   "ALARM_PT402" := ("PT402_VAL" > "PT402_HIGH") OR ("ALARM_PT402" AND NOT #CLEAR);
   "ALARM_PT501" := ("PT501_VAL" < "PT501_LOW_C") OR ("ALARM_PT501" AND NOT #CLEAR);
   "ALARM_PT502" := ("PT502_VAL" > "PT502_HIGH") OR ("ALARM_PT502" AND NOT #CLEAR);
   "ALARM_PT601" := ("PT601_VAL" >= "PT601_HIGH") OR ("ALARM_PT601" AND NOT #CLEAR);
   "ALARM_PT801" := ("PT801_VAL" < "PT801_LOW") OR ("ALARM_PT801" AND NOT #CLEAR);
   "ALARM_PT901" := ("PT901_VAL" > "PT901_HIGH") OR ("ALARM_PT901" AND NOT #CLEAR);
   "ALARM_DOORS_OPEN" := NOT "ABORT_ON" AND NOT "STEP_0_ON" AND NOT "DOORS_CLOSED" AND "AlwaysFALSE";
END_REGION

REGION Network 2
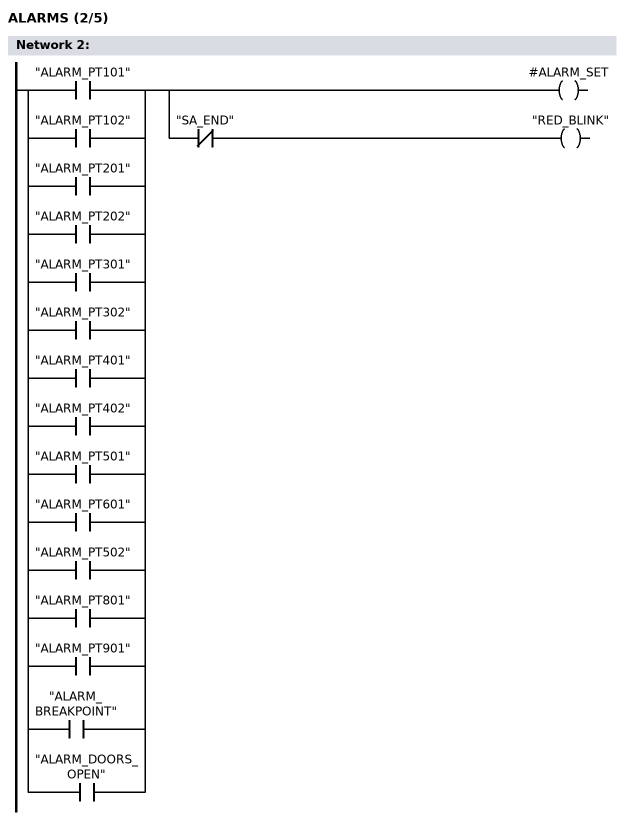
   RUNG wire#powerrail
      Contact( "ALARM_PT101" )
      wire#w1
      Coil( #ALARM_SET )
   END_RUNG
   RUNG wire#powerrail
      Contact( "ALARM_PT102" )
   END_RUNG wire#w1
   RUNG wire#powerrail
      Contact( "ALARM_PT201" )
   END_RUNG wire#w1
   RUNG wire#powerrail
      Contact( "ALARM_PT202" )
   END_RUNG wire#w1
   RUNG wire#powerrail
      Contact( "ALARM_PT301" )
   END_RUNG wire#w1
   RUNG wire#powerrail
      Contact( "ALARM_PT302" )
   END_RUNG wire#w1
   RUNG wire#powerrail
      Contact( "ALARM_PT401" )
   END_RUNG wire#w1
   RUNG wire#powerrail
      Contact( "ALARM_PT402" )
   END_RUNG wire#w1
   RUNG wire#powerrail
      Contact( "ALARM_PT501" )
   END_RUNG wire#w1
   RUNG wire#powerrail
      Contact( "ALARM_PT601" )
   END_RUNG wire#w1
   RUNG wire#powerrail
      Contact( "ALARM_PT502" )
   END_RUNG wire#w1
   RUNG wire#powerrail
      Contact( "ALARM_PT801" )
   END_RUNG wire#w1
   RUNG wire#powerrail
      Contact( "ALARM_PT901" )
   END_RUNG wire#w1
   RUNG wire#powerrail
      Contact( "ALARM_BREAKPOINT" )
   END_RUNG wire#w1
   RUNG wire#powerrail
      Contact( "ALARM_DOORS_OPEN" )
   END_RUNG wire#w1
   RUNG wire#w1
      I_Contact( "SA_END" )
      Coil( "RED_BLINK" )
   END_RUNG
   // the same network as SCL:
   #ALARM_SET := "ALARM_PT101" OR "ALARM_PT102" OR "ALARM_PT201" OR "ALARM_PT202" OR "ALARM_PT301" OR "ALARM_PT302" OR "ALARM_PT401" OR "ALARM_PT402" OR "ALARM_PT501" OR "ALARM_PT601" OR "ALARM_PT502" OR "ALARM_PT801" OR "ALARM_PT901" OR "ALARM_BREAKPOINT" OR "ALARM_DOORS_OPEN";
   "RED_BLINK" := #ALARM_SET AND NOT "SA_END";
END_REGION

REGION Network 3
   // PV701 Limit Switch Alarm
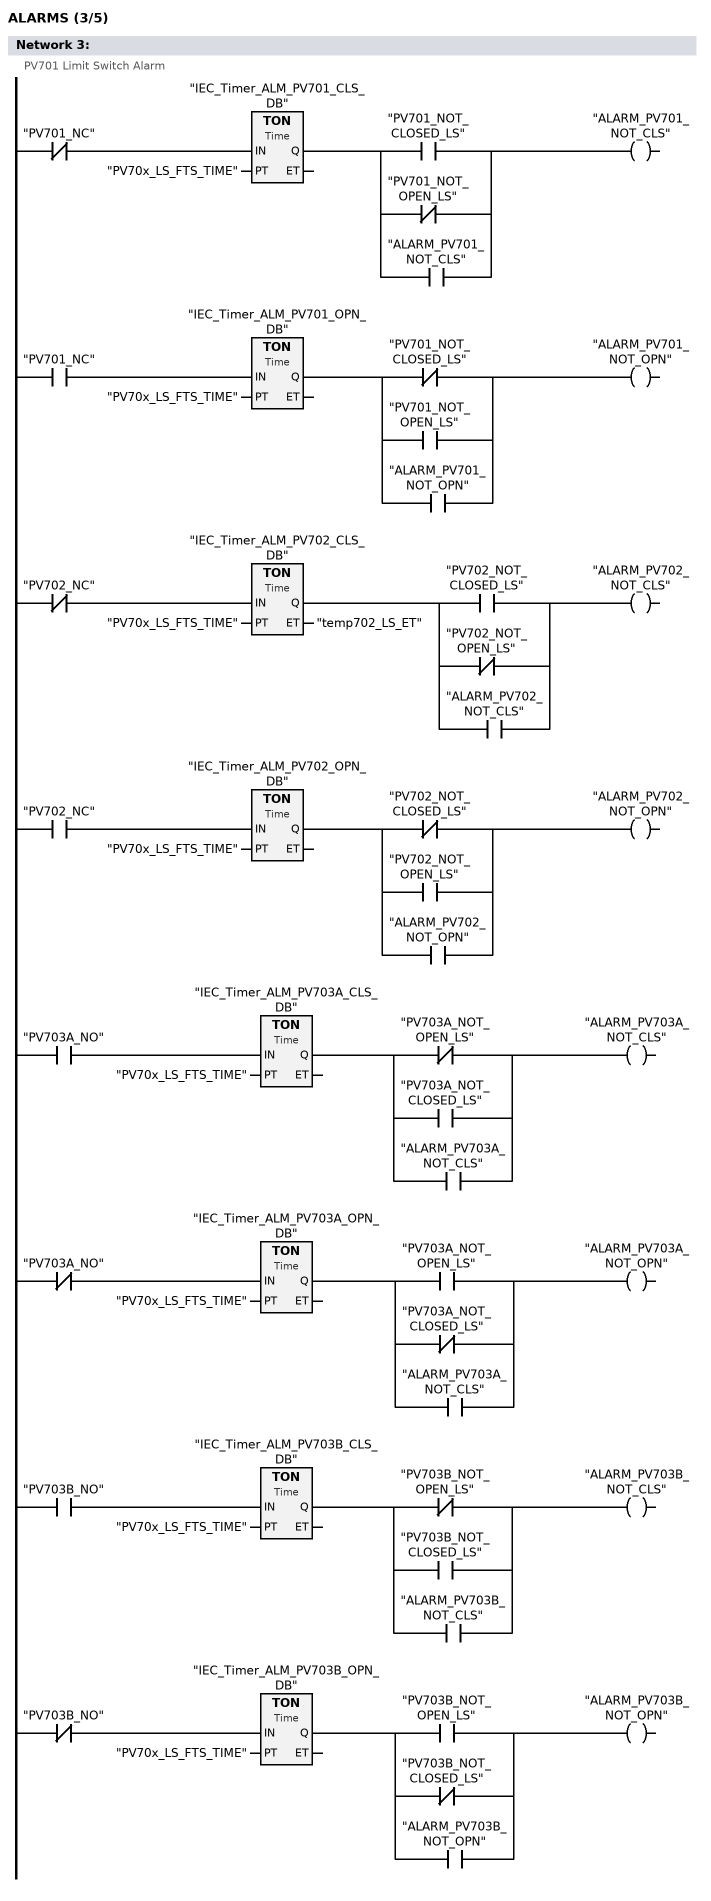
   "IEC_Timer_ALM_PV701_CLS_DB".TON(IN := NOT "PV701_NC", PT := "PV70x_LS_FTS_TIME");
   "ALARM_PV701_NOT_CLS" := "IEC_Timer_ALM_PV701_CLS_DB".Q AND ("PV701_NOT_CLOSED_LS" OR NOT "PV701_NOT_OPEN_LS" OR "ALARM_PV701_NOT_CLS");
   "IEC_Timer_ALM_PV701_OPN_DB".TON(IN := "PV701_NC", PT := "PV70x_LS_FTS_TIME");
   "ALARM_PV701_NOT_OPN" := "IEC_Timer_ALM_PV701_OPN_DB".Q AND (NOT "PV701_NOT_CLOSED_LS" OR "PV701_NOT_OPEN_LS" OR "ALARM_PV701_NOT_OPN");
   "IEC_Timer_ALM_PV702_CLS_DB".TON(IN := NOT "PV702_NC", PT := "PV70x_LS_FTS_TIME", ET => "temp702_LS_ET");
   "ALARM_PV702_NOT_CLS" := "IEC_Timer_ALM_PV702_CLS_DB".Q AND ("PV702_NOT_CLOSED_LS" OR NOT "PV702_NOT_OPEN_LS" OR "ALARM_PV702_NOT_CLS");
   "IEC_Timer_ALM_PV702_OPN_DB".TON(IN := "PV702_NC", PT := "PV70x_LS_FTS_TIME");
   "ALARM_PV702_NOT_OPN" := "IEC_Timer_ALM_PV702_OPN_DB".Q AND (NOT "PV702_NOT_CLOSED_LS" OR "PV702_NOT_OPEN_LS" OR "ALARM_PV702_NOT_OPN");
   "IEC_Timer_ALM_PV703A_CLS_DB".TON(IN := "PV703A_NO", PT := "PV70x_LS_FTS_TIME");
   "ALARM_PV703A_NOT_CLS" := "IEC_Timer_ALM_PV703A_CLS_DB".Q AND (NOT "PV703A_NOT_OPEN_LS" OR "PV703A_NOT_CLOSED_LS" OR "ALARM_PV703A_NOT_CLS");
   "IEC_Timer_ALM_PV703A_OPN_DB".TON(IN := NOT "PV703A_NO", PT := "PV70x_LS_FTS_TIME");
   "ALARM_PV703A_NOT_OPN" := "IEC_Timer_ALM_PV703A_OPN_DB".Q AND ("PV703A_NOT_OPEN_LS" OR NOT "PV703A_NOT_CLOSED_LS" OR "ALARM_PV703A_NOT_CLS");
   "IEC_Timer_ALM_PV703B_CLS_DB".TON(IN := "PV703B_NO", PT := "PV70x_LS_FTS_TIME");
   "ALARM_PV703B_NOT_CLS" := "IEC_Timer_ALM_PV703B_CLS_DB".Q AND (NOT "PV703B_NOT_OPEN_LS" OR "PV703B_NOT_CLOSED_LS" OR "ALARM_PV703B_NOT_CLS");
   "IEC_Timer_ALM_PV703B_OPN_DB".TON(IN := NOT "PV703B_NO", PT := "PV70x_LS_FTS_TIME");
   "ALARM_PV703B_NOT_OPN" := "IEC_Timer_ALM_PV703B_OPN_DB".Q AND ("PV703B_NOT_OPEN_LS" OR NOT "PV703B_NOT_CLOSED_LS" OR "ALARM_PV703B_NOT_OPN");
END_REGION

REGION Network 4
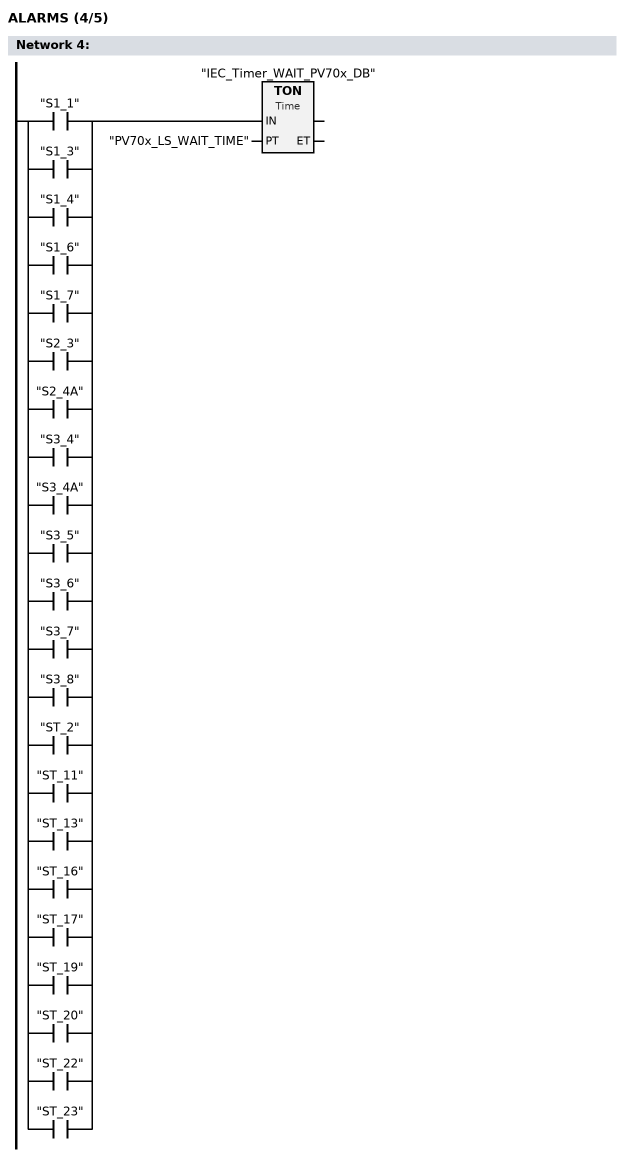
   "IEC_Timer_WAIT_PV70x_DB".TON(IN := "S1_1" OR "S1_3" OR "S1_4" OR "S1_6" OR "S1_7" OR "S2_3" OR "S2_4A" OR "S3_4" OR "S3_4A" OR "S3_5" OR "S3_6" OR "S3_7" OR "S3_8" OR "ST_2" OR "ST_11" OR "ST_13" OR "ST_16" OR "ST_17" OR "ST_19" OR "ST_20" OR "ST_22" OR "ST_23",
                           PT := "PV70x_LS_WAIT_TIME");
END_REGION

REGION Network 5
   // LIGHTS
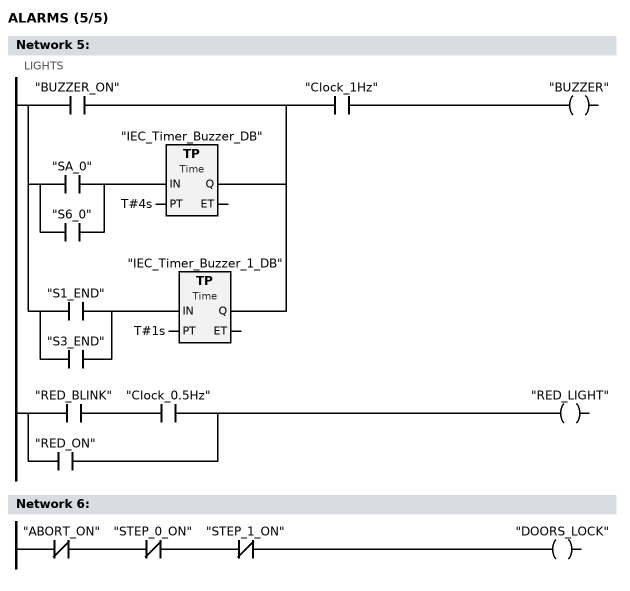
   "IEC_Timer_Buzzer_DB".TP(IN := "SA_0" OR "S6_0", PT := T#4s);
   "IEC_Timer_Buzzer_1_DB".TP(IN := "S1_END" OR "S3_END", PT := T#1s);
   "BUZZER" := ("BUZZER_ON" OR "IEC_Timer_Buzzer_DB".Q OR "IEC_Timer_Buzzer_1_DB".Q) AND "Clock_1Hz";
   "RED_LIGHT" := ("RED_BLINK" AND "Clock_0.5Hz") OR "RED_ON";
END_REGION

REGION Network 6
   RUNG wire#powerrail
      I_Contact( "ABORT_ON" )
      I_Contact( "STEP_0_ON" )
      I_Contact( "STEP_1_ON" )
      Coil( "DOORS_LOCK" )
   END_RUNG
   // the same network as SCL:
   "DOORS_LOCK" := NOT "ABORT_ON" AND NOT "STEP_0_ON" AND NOT "STEP_1_ON";
END_REGION
END_FUNCTION

FUNCTION "ABORTING" : Void   // FC15, LAD
{ S7_Optimized_Access := 'FALSE' }
VERSION : 0.1
// Modified to Fully open MFC601
BEGIN

REGION Network 2
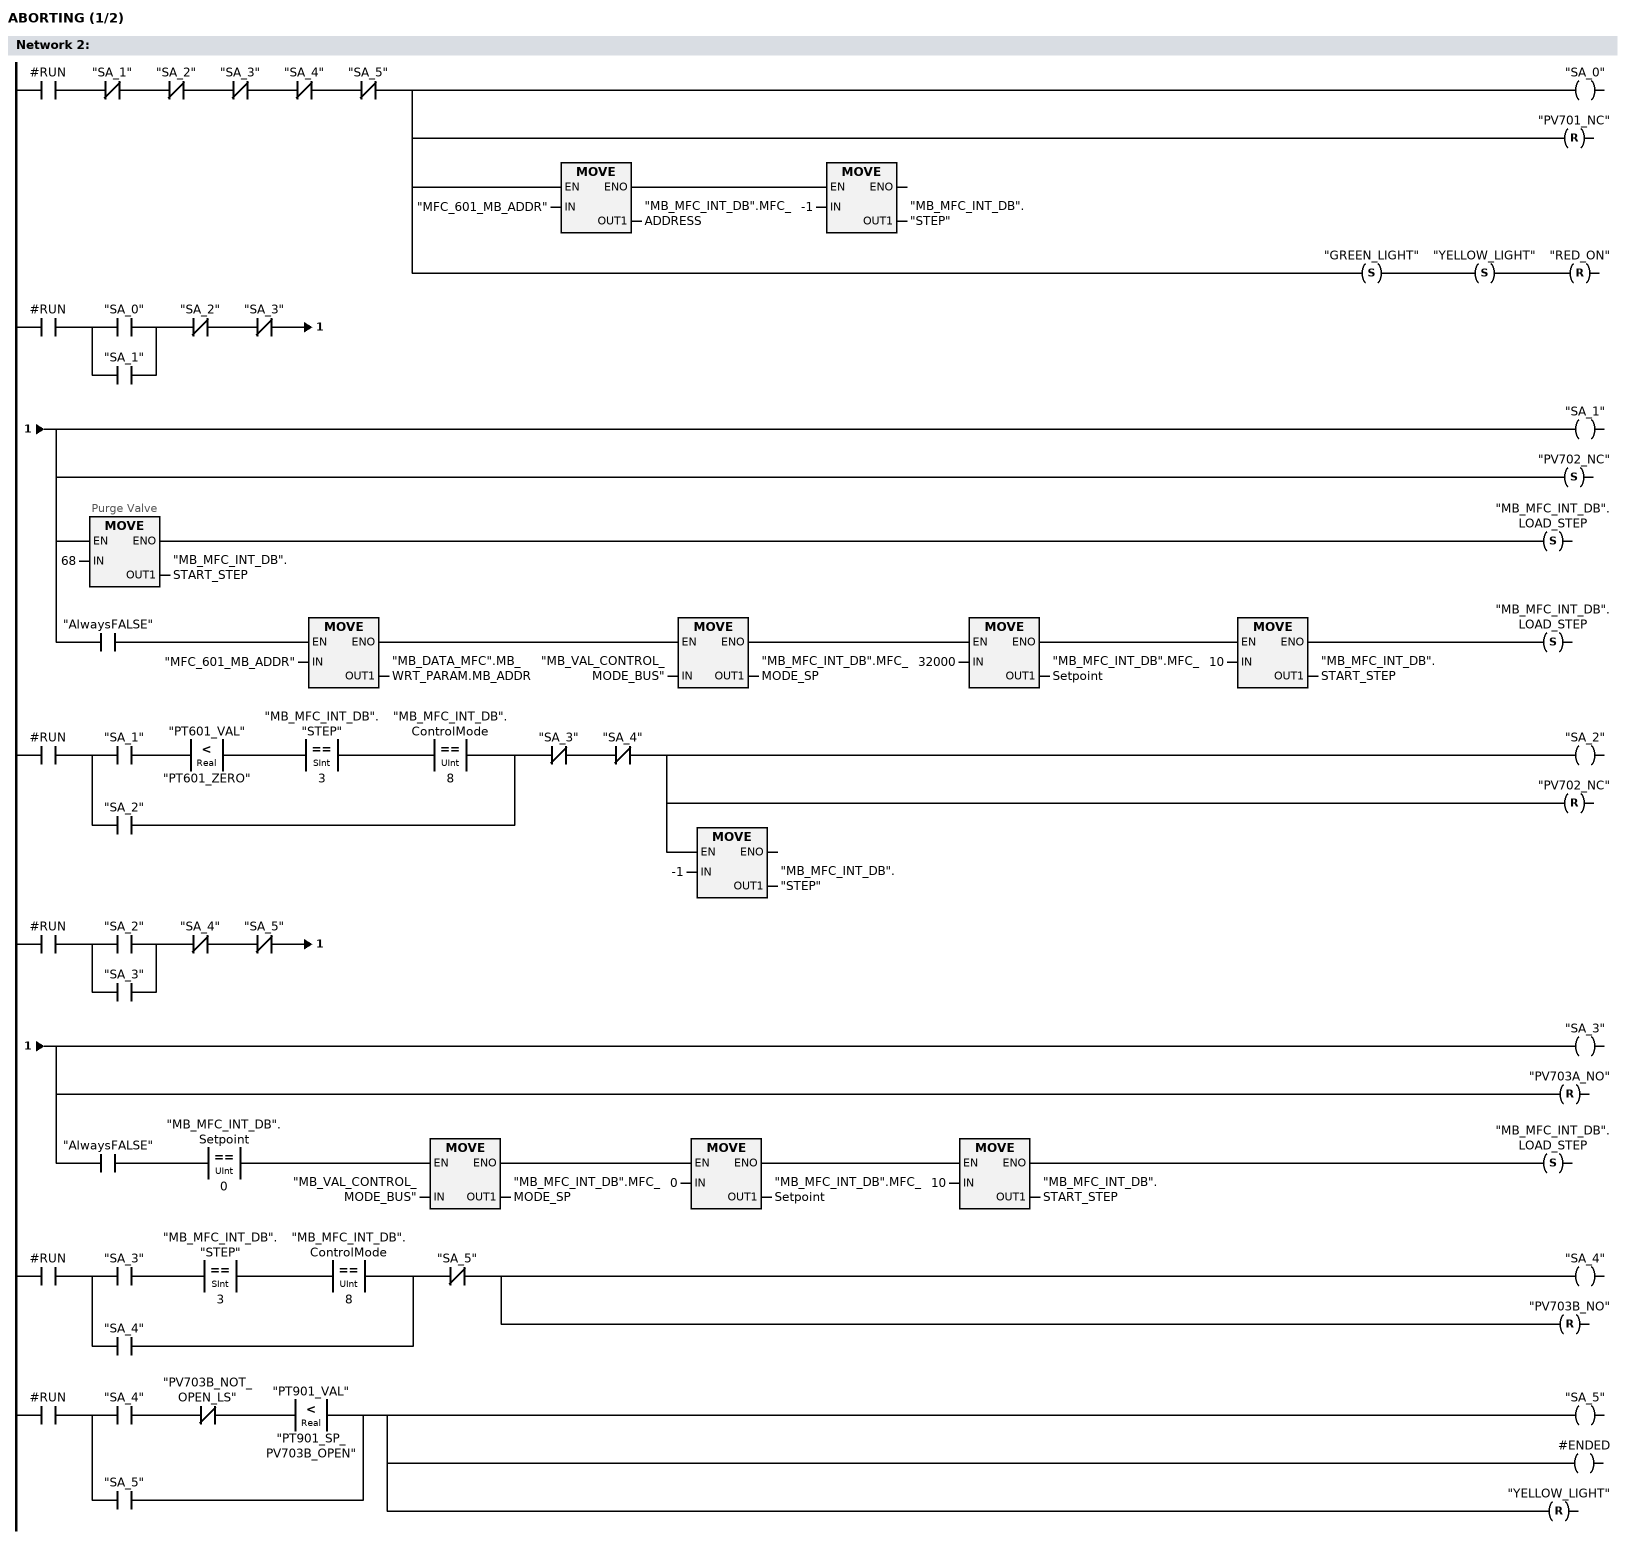
   RUNG wire#powerrail
      Contact( #RUN )
      I_Contact( "SA_1" )
      I_Contact( "SA_2" )
      I_Contact( "SA_3" )
      I_Contact( "SA_4" )
      I_Contact( "SA_5" )
      wire#w1
      Coil( "SA_0" )
   END_RUNG
   RUNG wire#w1
      R_Coil( "PV701_NC" )
   END_RUNG
   RUNG wire#w1
      Move(in := "MFC_601_MB_ADDR", out1 => "MB_MFC_INT_DB".MFC_ADDRESS)
      Move(in := -1, out1 => "MB_MFC_INT_DB"."STEP")
   END_RUNG
   RUNG wire#w1
      S_Coil( "GREEN_LIGHT" )
      S_Coil( "YELLOW_LIGHT" )
      R_Coil( "RED_ON" )
   END_RUNG
   RUNG wire#powerrail
      Contact( #RUN )
      wire#w2
      Contact( "SA_0" )
      wire#w3
      I_Contact( "SA_2" )
      I_Contact( "SA_3" )
      wire#w4
      Coil( "SA_1" )
   END_RUNG
   RUNG wire#w2
      Contact( "SA_1" )
   END_RUNG wire#w3
   RUNG wire#w4
      S_Coil( "PV702_NC" )
   END_RUNG
   RUNG wire#w4
      Move(in := 68, out1 => "MB_MFC_INT_DB".START_STEP)   // Purge Valve
      S_Coil( "MB_MFC_INT_DB".LOAD_STEP )
   END_RUNG
   RUNG wire#w4
      Contact( "AlwaysFALSE" )
      Move(in := "MFC_601_MB_ADDR", out1 => "MB_DATA_MFC".MB_WRT_PARAM.MB_ADDR)
      Move(in := "MB_VAL_CONTROL_MODE_BUS", out1 => "MB_MFC_INT_DB".MFC_MODE_SP)
      Move(in := 32000, out1 => "MB_MFC_INT_DB".MFC_Setpoint)
      Move(in := 10, out1 => "MB_MFC_INT_DB".START_STEP)
      S_Coil( "MB_MFC_INT_DB".LOAD_STEP )
   END_RUNG
   RUNG wire#powerrail
      Contact( #RUN )
      wire#w5
      Contact( "SA_1" )
      { S7_Templates := "SrcType := Real" } LT_Contact(in1 := "PT601_VAL", in2 := "PT601_ZERO")
      { S7_Templates := "SrcType := SInt" } EQ_Contact(in1 := "MB_MFC_INT_DB"."STEP", in2 := 3)
      { S7_Templates := "SrcType := UInt" } EQ_Contact(in1 := "MB_MFC_INT_DB".ControlMode, in2 := 8)
      wire#w6
      I_Contact( "SA_3" )
      I_Contact( "SA_4" )
      wire#w7
      Coil( "SA_2" )
   END_RUNG
   RUNG wire#w5
      Contact( "SA_2" )
   END_RUNG wire#w6
   RUNG wire#w7
      R_Coil( "PV702_NC" )
   END_RUNG
   RUNG wire#w7
      Move(in := -1, out1 => "MB_MFC_INT_DB"."STEP")
   END_RUNG
   RUNG wire#powerrail
      Contact( #RUN )
      wire#w8
      Contact( "SA_2" )
      wire#w9
      I_Contact( "SA_4" )
      I_Contact( "SA_5" )
      wire#w10
      Coil( "SA_3" )
   END_RUNG
   RUNG wire#w8
      Contact( "SA_3" )
   END_RUNG wire#w9
   RUNG wire#w10
      R_Coil( "PV703A_NO" )
   END_RUNG
   RUNG wire#w10
      Contact( "AlwaysFALSE" )
      { S7_Templates := "SrcType := UInt" } EQ_Contact(in1 := "MB_MFC_INT_DB".Setpoint, in2 := 0)
      Move(in := "MB_VAL_CONTROL_MODE_BUS", out1 => "MB_MFC_INT_DB".MFC_MODE_SP)
      Move(in := 0, out1 => "MB_MFC_INT_DB".MFC_Setpoint)
      Move(in := 10, out1 => "MB_MFC_INT_DB".START_STEP)
      S_Coil( "MB_MFC_INT_DB".LOAD_STEP )
   END_RUNG
   RUNG wire#powerrail
      Contact( #RUN )
      wire#w11
      Contact( "SA_3" )
      { S7_Templates := "SrcType := SInt" } EQ_Contact(in1 := "MB_MFC_INT_DB"."STEP", in2 := 3)
      { S7_Templates := "SrcType := UInt" } EQ_Contact(in1 := "MB_MFC_INT_DB".ControlMode, in2 := 8)
      wire#w12
      I_Contact( "SA_5" )
      wire#w13
      Coil( "SA_4" )
   END_RUNG
   RUNG wire#w11
      Contact( "SA_4" )
   END_RUNG wire#w12
   RUNG wire#w13
      R_Coil( "PV703B_NO" )
   END_RUNG
   RUNG wire#powerrail
      Contact( #RUN )
      wire#w14
      Contact( "SA_4" )
      I_Contact( "PV703B_NOT_OPEN_LS" )
      { S7_Templates := "SrcType := Real" } LT_Contact(in1 := "PT901_VAL", in2 := "PT901_SP_PV703B_OPEN")
      wire#w15
      Coil( "SA_5" )
   END_RUNG
   RUNG wire#w14
      Contact( "SA_5" )
   END_RUNG wire#w15
   RUNG wire#w15
      Coil( #ENDED )
   END_RUNG
   RUNG wire#w15
      R_Coil( "YELLOW_LIGHT" )
   END_RUNG
   // the same network as SCL:
   "SA_0" := #RUN AND NOT "SA_1" AND NOT "SA_2" AND NOT "SA_3" AND NOT "SA_4" AND NOT "SA_5";
   IF "SA_0" THEN
       "PV701_NC" := FALSE;
       "MB_MFC_INT_DB".MFC_ADDRESS := "MFC_601_MB_ADDR";
       "MB_MFC_INT_DB"."STEP" := -1;
       "GREEN_LIGHT" := TRUE;
       "YELLOW_LIGHT" := TRUE;
       "RED_ON" := FALSE;
   END_IF;
   "SA_1" := #RUN AND ("SA_0" OR "SA_1") AND NOT "SA_2" AND NOT "SA_3";
   IF "SA_1" THEN
       "PV702_NC" := TRUE;
       "MB_MFC_INT_DB".START_STEP := 68;   // Purge Valve
       "MB_MFC_INT_DB".LOAD_STEP := TRUE;
   END_IF;
   IF "SA_1" AND "AlwaysFALSE" THEN
       "MB_DATA_MFC".MB_WRT_PARAM.MB_ADDR := "MFC_601_MB_ADDR";
       "MB_MFC_INT_DB".MFC_MODE_SP := "MB_VAL_CONTROL_MODE_BUS";
       "MB_MFC_INT_DB".MFC_Setpoint := 32000;
       "MB_MFC_INT_DB".START_STEP := 10;
       "MB_MFC_INT_DB".LOAD_STEP := TRUE;
   END_IF;
   "SA_2" := #RUN AND (("SA_1" AND ("PT601_VAL" < "PT601_ZERO") AND ("MB_MFC_INT_DB"."STEP" = 3) AND ("MB_MFC_INT_DB".ControlMode = 8)) OR "SA_2") AND NOT "SA_3" AND NOT "SA_4";
   IF "SA_2" THEN
       "PV702_NC" := FALSE;
       "MB_MFC_INT_DB"."STEP" := -1;
   END_IF;
   "SA_3" := #RUN AND ("SA_2" OR "SA_3") AND NOT "SA_4" AND NOT "SA_5";
   IF "SA_3" THEN "PV703A_NO" := FALSE; END_IF;
   IF "SA_3" AND "AlwaysFALSE" AND ("MB_MFC_INT_DB".Setpoint = 0) THEN
       "MB_MFC_INT_DB".MFC_MODE_SP := "MB_VAL_CONTROL_MODE_BUS";
       "MB_MFC_INT_DB".MFC_Setpoint := 0;
       "MB_MFC_INT_DB".START_STEP := 10;
       "MB_MFC_INT_DB".LOAD_STEP := TRUE;
   END_IF;
   "SA_4" := #RUN AND (("SA_3" AND ("MB_MFC_INT_DB"."STEP" = 3) AND ("MB_MFC_INT_DB".ControlMode = 8)) OR "SA_4") AND NOT "SA_5";
   IF "SA_4" THEN "PV703B_NO" := FALSE; END_IF;
   "SA_5" := #RUN AND (("SA_4" AND NOT "PV703B_NOT_OPEN_LS" AND ("PT901_VAL" < "PT901_SP_PV703B_OPEN")) OR "SA_5");
   #ENDED := "SA_5";
   IF "SA_5" THEN "YELLOW_LIGHT" := FALSE; END_IF;
END_REGION

REGION Network 3: NC
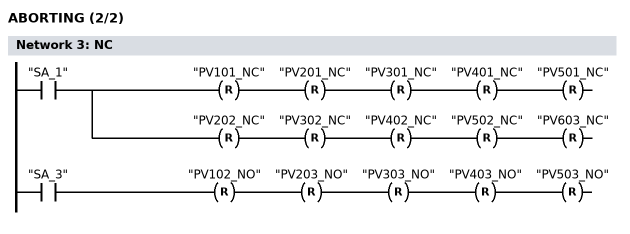
   RUNG wire#powerrail
      Contact( "SA_1" )
      wire#w1
      R_Coil( "PV101_NC" )
      R_Coil( "PV201_NC" )
      R_Coil( "PV301_NC" )
      R_Coil( "PV401_NC" )
      R_Coil( "PV501_NC" )
   END_RUNG
   RUNG wire#w1
      R_Coil( "PV202_NC" )
      R_Coil( "PV302_NC" )
      R_Coil( "PV402_NC" )
      R_Coil( "PV502_NC" )
      R_Coil( "PV603_NC" )
   END_RUNG
   RUNG wire#powerrail
      Contact( "SA_3" )
      R_Coil( "PV102_NO" )
      R_Coil( "PV203_NO" )
      R_Coil( "PV303_NO" )
      R_Coil( "PV403_NO" )
      R_Coil( "PV503_NO" )
   END_RUNG
   // the same network as SCL:
   IF "SA_1" THEN
       "PV101_NC" := FALSE;
       "PV201_NC" := FALSE;
       "PV301_NC" := FALSE;
       "PV401_NC" := FALSE;
       "PV501_NC" := FALSE;
       "PV202_NC" := FALSE;
       "PV302_NC" := FALSE;
       "PV402_NC" := FALSE;
       "PV502_NC" := FALSE;
       "PV603_NC" := FALSE;
   END_IF;
   IF "SA_3" THEN
       "PV102_NO" := FALSE;
       "PV203_NO" := FALSE;
       "PV303_NO" := FALSE;
       "PV403_NO" := FALSE;
       "PV503_NO" := FALSE;
   END_IF;
END_REGION
END_FUNCTION

FUNCTION "ALL_VALVES_STANDBY" : Void   // FC16, LAD
{ S7_Optimized_Access := 'FALSE' }
VERSION : 0.1
// All Valves on Stant by Mode
BEGIN

REGION Network 1: NC
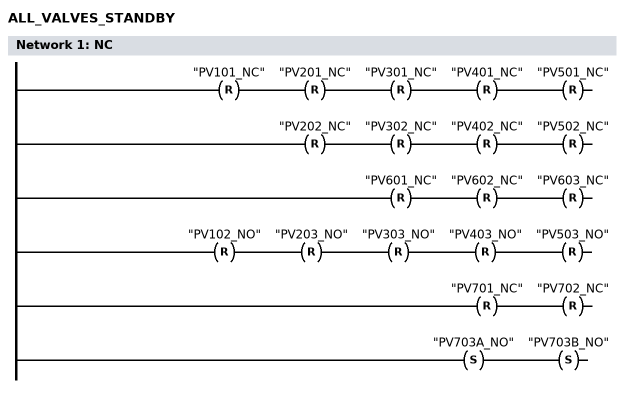
   RUNG wire#powerrail
      R_Coil( "PV101_NC" )
      R_Coil( "PV201_NC" )
      R_Coil( "PV301_NC" )
      R_Coil( "PV401_NC" )
      R_Coil( "PV501_NC" )
   END_RUNG
   RUNG wire#powerrail
      R_Coil( "PV202_NC" )
      R_Coil( "PV302_NC" )
      R_Coil( "PV402_NC" )
      R_Coil( "PV502_NC" )
   END_RUNG
   RUNG wire#powerrail
      R_Coil( "PV601_NC" )
      R_Coil( "PV602_NC" )
      R_Coil( "PV603_NC" )
   END_RUNG
   RUNG wire#powerrail
      R_Coil( "PV102_NO" )
      R_Coil( "PV203_NO" )
      R_Coil( "PV303_NO" )
      R_Coil( "PV403_NO" )
      R_Coil( "PV503_NO" )
   END_RUNG
   RUNG wire#powerrail
      R_Coil( "PV701_NC" )
      R_Coil( "PV702_NC" )
   END_RUNG
   RUNG wire#powerrail
      S_Coil( "PV703A_NO" )
      S_Coil( "PV703B_NO" )
   END_RUNG
   // the same network as SCL:
   "PV101_NC" := FALSE;
   "PV201_NC" := FALSE;
   "PV301_NC" := FALSE;
   "PV401_NC" := FALSE;
   "PV501_NC" := FALSE;
   "PV202_NC" := FALSE;
   "PV302_NC" := FALSE;
   "PV402_NC" := FALSE;
   "PV502_NC" := FALSE;
   "PV601_NC" := FALSE;
   "PV602_NC" := FALSE;
   "PV603_NC" := FALSE;
   "PV102_NO" := FALSE;
   "PV203_NO" := FALSE;
   "PV303_NO" := FALSE;
   "PV403_NO" := FALSE;
   "PV503_NO" := FALSE;
   "PV701_NC" := FALSE;
   "PV702_NC" := FALSE;
   "PV703A_NO" := TRUE;
   "PV703B_NO" := TRUE;
END_REGION
END_FUNCTION

FUNCTION "TESTS_3" : Void   // FC17, LAD
{ S7_Optimized_Access := 'FALSE' }
VERSION : 0.1
// Test_MFC601
   VAR_TEMP   // added for the SCL form of the ladder/FBD networks
      _w1 : Bool;
   END_VAR
BEGIN

REGION Network 1
   // ALARM Settings
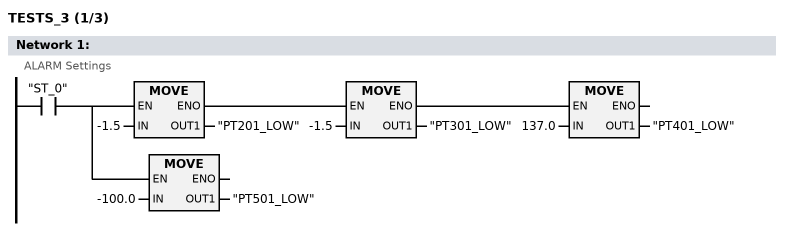
   RUNG wire#powerrail
      Contact( "ST_0" )
      wire#w1
      { S7_GenerateENO := "TRUE" } Move(in := -1.5, out1 => "PT201_LOW")
      { S7_GenerateENO := "TRUE" } Move(in := -1.5, out1 => "PT301_LOW")
      { S7_GenerateENO := "TRUE" } Move(in := 137.0, out1 => "PT401_LOW")
   END_RUNG
   RUNG wire#w1
      { S7_GenerateENO := "TRUE" } Move(in := -100.0, out1 => "PT501_LOW")
   END_RUNG
   // the same network as SCL:
   // ENO of a box is taken as its EN; it also drops when the box reports an error
   IF "ST_0" THEN
       "PT201_LOW" := -1.5;
       "PT301_LOW" := -1.5;
       "PT401_LOW" := 137.0;
       "PT501_LOW" := -100.0;
   END_IF;
END_REGION

REGION Network 2: Pneumatic Tests
   // Test Pneumatic System (Test #1-#6)
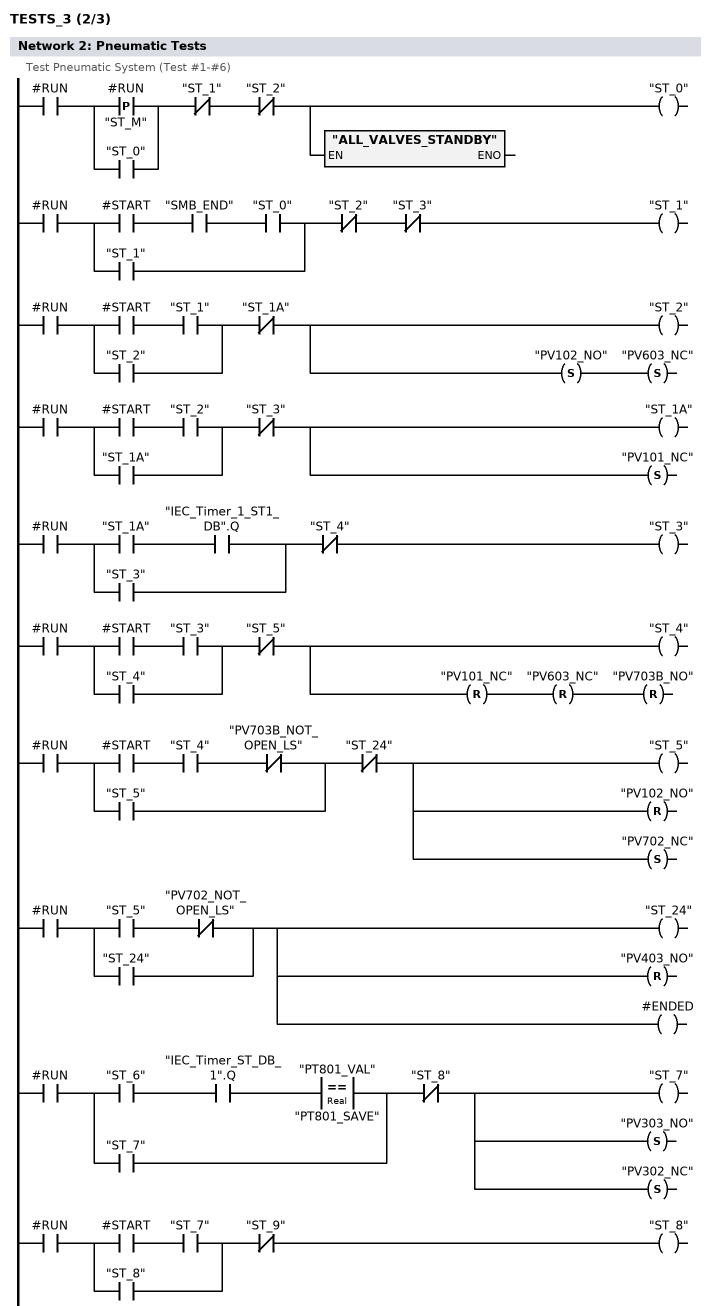
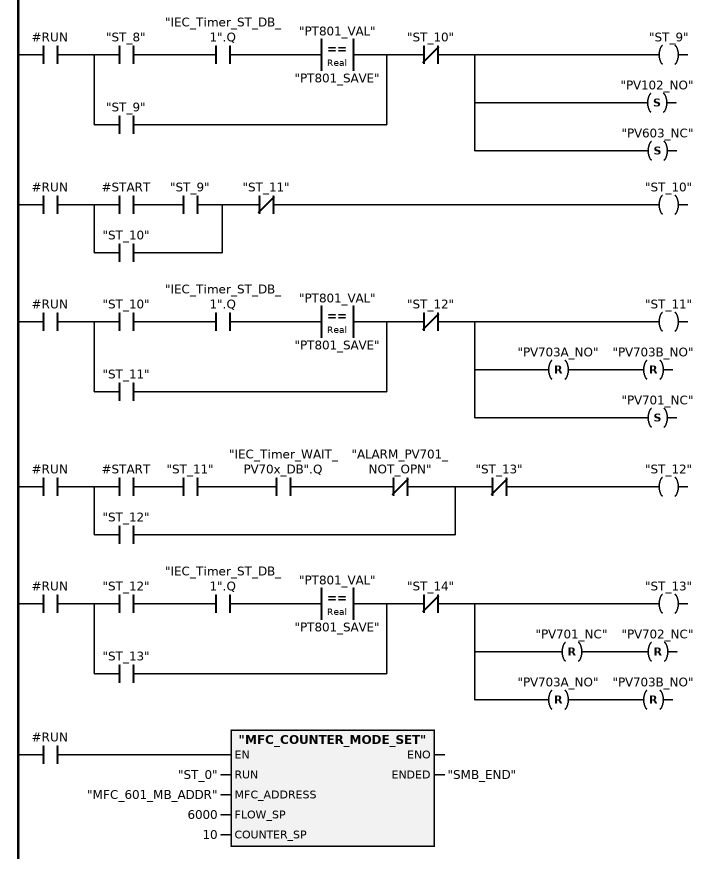
   RUNG wire#powerrail
      Contact( #RUN )
      wire#w1
      P_Contact(operand := #RUN, bit := "ST_M")
      wire#w2
      I_Contact( "ST_1" )
      I_Contact( "ST_2" )
      wire#w3
      Coil( "ST_0" )
   END_RUNG
   RUNG wire#w1
      Contact( "ST_0" )
   END_RUNG wire#w2
   RUNG wire#w3
      "ALL_VALVES_STANDBY"()
   END_RUNG
   RUNG wire#powerrail
      Contact( #RUN )
      wire#w4
      Contact( #START )
      Contact( "SMB_END" )
      Contact( "ST_0" )
      wire#w5
      I_Contact( "ST_2" )
      I_Contact( "ST_3" )
      Coil( "ST_1" )
   END_RUNG
   RUNG wire#w4
      Contact( "ST_1" )
   END_RUNG wire#w5
   RUNG wire#powerrail
      Contact( #RUN )
      wire#w6
      Contact( #START )
      Contact( "ST_1" )
      wire#w7
      I_Contact( "ST_1A" )
      wire#w8
      Coil( "ST_2" )
   END_RUNG
   RUNG wire#w6
      Contact( "ST_2" )
   END_RUNG wire#w7
   RUNG wire#w8
      S_Coil( "PV102_NO" )
      S_Coil( "PV603_NC" )
   END_RUNG
   RUNG wire#powerrail
      Contact( #RUN )
      wire#w9
      Contact( #START )
      Contact( "ST_2" )
      wire#w10
      I_Contact( "ST_3" )
      wire#w11
      Coil( "ST_1A" )
   END_RUNG
   RUNG wire#w9
      Contact( "ST_1A" )
   END_RUNG wire#w10
   RUNG wire#w11
      S_Coil( "PV101_NC" )
   END_RUNG
   RUNG wire#powerrail
      Contact( #RUN )
      wire#w12
      Contact( "ST_1A" )
      Contact( "IEC_Timer_1_ST1_DB".Q )
      wire#w13
      I_Contact( "ST_4" )
      Coil( "ST_3" )
   END_RUNG
   RUNG wire#w12
      Contact( "ST_3" )
   END_RUNG wire#w13
   RUNG wire#powerrail
      Contact( #RUN )
      wire#w14
      Contact( #START )
      Contact( "ST_3" )
      wire#w15
      I_Contact( "ST_5" )
      wire#w16
      Coil( "ST_4" )
   END_RUNG
   RUNG wire#w14
      Contact( "ST_4" )
   END_RUNG wire#w15
   RUNG wire#w16
      R_Coil( "PV101_NC" )
      R_Coil( "PV603_NC" )
      R_Coil( "PV703B_NO" )
   END_RUNG
   RUNG wire#powerrail
      Contact( #RUN )
      wire#w17
      Contact( #START )
      Contact( "ST_4" )
      I_Contact( "PV703B_NOT_OPEN_LS" )
      wire#w18
      I_Contact( "ST_24" )
      wire#w19
      Coil( "ST_5" )
   END_RUNG
   RUNG wire#w17
      Contact( "ST_5" )
   END_RUNG wire#w18
   RUNG wire#w19
      R_Coil( "PV102_NO" )
   END_RUNG
   RUNG wire#w19
      S_Coil( "PV702_NC" )
   END_RUNG
   RUNG wire#powerrail
      Contact( #RUN )
      wire#w20
      Contact( "ST_5" )
      I_Contact( "PV702_NOT_OPEN_LS" )
      wire#w21
      Coil( "ST_24" )
   END_RUNG
   RUNG wire#w20
      Contact( "ST_24" )
   END_RUNG wire#w21
   RUNG wire#w21
      R_Coil( "PV403_NO" )
   END_RUNG
   RUNG wire#w21
      Coil( #ENDED )
   END_RUNG
   RUNG wire#powerrail
      Contact( #RUN )
      wire#w22
      Contact( "ST_6" )
      Contact( "IEC_Timer_ST_DB_1".Q )
      { S7_Templates := "SrcType := Real" } EQ_Contact(in1 := "PT801_VAL", in2 := "PT801_SAVE")
      wire#w23
      I_Contact( "ST_8" )
      wire#w24
      Coil( "ST_7" )
   END_RUNG
   RUNG wire#w22
      Contact( "ST_7" )
   END_RUNG wire#w23
   RUNG wire#w24
      S_Coil( "PV303_NO" )
   END_RUNG
   RUNG wire#w24
      S_Coil( "PV302_NC" )
   END_RUNG
   RUNG wire#powerrail
      Contact( #RUN )
      wire#w25
      Contact( #START )
      Contact( "ST_7" )
      wire#w26
      I_Contact( "ST_9" )
      Coil( "ST_8" )
   END_RUNG
   RUNG wire#w25
      Contact( "ST_8" )
   END_RUNG wire#w26
   RUNG wire#powerrail
      Contact( #RUN )
      wire#w27
      Contact( "ST_8" )
      Contact( "IEC_Timer_ST_DB_1".Q )
      { S7_Templates := "SrcType := Real" } EQ_Contact(in1 := "PT801_VAL", in2 := "PT801_SAVE")
      wire#w28
      I_Contact( "ST_10" )
      wire#w29
      Coil( "ST_9" )
   END_RUNG
   RUNG wire#w27
      Contact( "ST_9" )
   END_RUNG wire#w28
   RUNG wire#w29
      S_Coil( "PV102_NO" )
   END_RUNG
   RUNG wire#w29
      S_Coil( "PV603_NC" )
   END_RUNG
   RUNG wire#powerrail
      Contact( #RUN )
      wire#w30
      Contact( #START )
      Contact( "ST_9" )
      wire#w31
      I_Contact( "ST_11" )
      Coil( "ST_10" )
   END_RUNG
   RUNG wire#w30
      Contact( "ST_10" )
   END_RUNG wire#w31
   RUNG wire#powerrail
      Contact( #RUN )
      wire#w32
      Contact( "ST_10" )
      Contact( "IEC_Timer_ST_DB_1".Q )
      { S7_Templates := "SrcType := Real" } EQ_Contact(in1 := "PT801_VAL", in2 := "PT801_SAVE")
      wire#w33
      I_Contact( "ST_12" )
      wire#w34
      Coil( "ST_11" )
   END_RUNG
   RUNG wire#w32
      Contact( "ST_11" )
   END_RUNG wire#w33
   RUNG wire#w34
      R_Coil( "PV703A_NO" )
      R_Coil( "PV703B_NO" )
   END_RUNG
   RUNG wire#w34
      S_Coil( "PV701_NC" )
   END_RUNG
   RUNG wire#powerrail
      Contact( #RUN )
      wire#w35
      Contact( #START )
      Contact( "ST_11" )
      Contact( "IEC_Timer_WAIT_PV70x_DB".Q )
      I_Contact( "ALARM_PV701_NOT_OPN" )
      wire#w36
      I_Contact( "ST_13" )
      Coil( "ST_12" )
   END_RUNG
   RUNG wire#w35
      Contact( "ST_12" )
   END_RUNG wire#w36
   RUNG wire#powerrail
      Contact( #RUN )
      wire#w37
      Contact( "ST_12" )
      Contact( "IEC_Timer_ST_DB_1".Q )
      { S7_Templates := "SrcType := Real" } EQ_Contact(in1 := "PT801_VAL", in2 := "PT801_SAVE")
      wire#w38
      I_Contact( "ST_14" )
      wire#w39
      Coil( "ST_13" )
   END_RUNG
   RUNG wire#w37
      Contact( "ST_13" )
   END_RUNG wire#w38
   RUNG wire#w39
      R_Coil( "PV701_NC" )
      R_Coil( "PV702_NC" )
   END_RUNG
   RUNG wire#w39
      R_Coil( "PV703A_NO" )
      R_Coil( "PV703B_NO" )
   END_RUNG
   RUNG wire#powerrail
      Contact( #RUN )
      "MFC_COUNTER_MODE_SET"(RUN := "ST_0", MFC_ADDRESS := "MFC_601_MB_ADDR", FLOW_SP := 6000, COUNTER_SP := 10, ENDED => "SMB_END")
   END_RUNG
   // the same network as SCL:
   #_w1 := #RUN AND #RUN AND NOT "ST_M";   // rising edge of #RUN
   "ST_M" := #RUN;
   "ST_0" := (#_w1 OR (#RUN AND "ST_0")) AND NOT "ST_1" AND NOT "ST_2";
   IF "ST_0" THEN "ALL_VALVES_STANDBY"(); END_IF;
   "ST_1" := #RUN AND ((#START AND "SMB_END" AND "ST_0") OR "ST_1") AND NOT "ST_2" AND NOT "ST_3";
   "ST_2" := #RUN AND ((#START AND "ST_1") OR "ST_2") AND NOT "ST_1A";
   IF "ST_2" THEN
       "PV102_NO" := TRUE;
       "PV603_NC" := TRUE;
   END_IF;
   "ST_1A" := #RUN AND ((#START AND "ST_2") OR "ST_1A") AND NOT "ST_3";
   IF "ST_1A" THEN "PV101_NC" := TRUE; END_IF;
   "ST_3" := #RUN AND (("ST_1A" AND "IEC_Timer_1_ST1_DB".Q) OR "ST_3") AND NOT "ST_4";
   "ST_4" := #RUN AND ((#START AND "ST_3") OR "ST_4") AND NOT "ST_5";
   IF "ST_4" THEN
       "PV101_NC" := FALSE;
       "PV603_NC" := FALSE;
       "PV703B_NO" := FALSE;
   END_IF;
   "ST_5" := #RUN AND ((#START AND "ST_4" AND NOT "PV703B_NOT_OPEN_LS") OR "ST_5") AND NOT "ST_24";
   IF "ST_5" THEN
       "PV102_NO" := FALSE;
       "PV702_NC" := TRUE;
   END_IF;
   "ST_24" := #RUN AND (("ST_5" AND NOT "PV702_NOT_OPEN_LS") OR "ST_24");
   IF "ST_24" THEN "PV403_NO" := FALSE; END_IF;
   #ENDED := "ST_24";
   "ST_7" := #RUN AND (("ST_6" AND "IEC_Timer_ST_DB_1".Q AND ("PT801_VAL" = "PT801_SAVE")) OR "ST_7") AND NOT "ST_8";
   IF "ST_7" THEN
       "PV303_NO" := TRUE;
       "PV302_NC" := TRUE;
   END_IF;
   "ST_8" := #RUN AND ((#START AND "ST_7") OR "ST_8") AND NOT "ST_9";
   "ST_9" := #RUN AND (("ST_8" AND "IEC_Timer_ST_DB_1".Q AND ("PT801_VAL" = "PT801_SAVE")) OR "ST_9") AND NOT "ST_10";
   IF "ST_9" THEN
       "PV102_NO" := TRUE;
       "PV603_NC" := TRUE;
   END_IF;
   "ST_10" := #RUN AND ((#START AND "ST_9") OR "ST_10") AND NOT "ST_11";
   "ST_11" := #RUN AND (("ST_10" AND "IEC_Timer_ST_DB_1".Q AND ("PT801_VAL" = "PT801_SAVE")) OR "ST_11") AND NOT "ST_12";
   IF "ST_11" THEN
       "PV703A_NO" := FALSE;
       "PV703B_NO" := FALSE;
       "PV701_NC" := TRUE;
   END_IF;
   "ST_12" := #RUN AND ((#START AND "ST_11" AND "IEC_Timer_WAIT_PV70x_DB".Q AND NOT "ALARM_PV701_NOT_OPN") OR "ST_12") AND NOT "ST_13";
   "ST_13" := #RUN AND (("ST_12" AND "IEC_Timer_ST_DB_1".Q AND ("PT801_VAL" = "PT801_SAVE")) OR "ST_13") AND NOT "ST_14";
   IF "ST_13" THEN
       "PV701_NC" := FALSE;
       "PV702_NC" := FALSE;
       "PV703A_NO" := FALSE;
       "PV703B_NO" := FALSE;
   END_IF;
   IF #RUN THEN
       "MFC_COUNTER_MODE_SET"(RUN := "ST_0",
                              MFC_ADDRESS := "MFC_601_MB_ADDR",
                              FLOW_SP := 6000,
                              COUNTER_SP := 10,
                              ENDED => "SMB_END");
   END_IF;
END_REGION

REGION Network 3: Process Tests
   // Tests Process Circuits  (Test #7-#9)
END_REGION

REGION Network 4
